REGION Network 96: "PALLET_PARA_ASCENSOR"
   RUNG wire#powerrail
      Contact( #Aux_1 )
      wire#w1
      Coil( "PALLET_PARA_ASCENSOR" )
   END_RUNG
   RUNG wire#powerrail
      Contact( "PALLET_PARA_ASCENSOR" )
      I_Contact( "Tonof_PALLET_EN_ASCENSOR" )
   END_RUNG wire#w1
   // the same network as SCL:
   "PALLET_PARA_ASCENSOR" := #Aux_1 OR ("PALLET_PARA_ASCENSOR" AND NOT "Tonof_PALLET_EN_ASCENSOR");
END_REGION

REGION Network 97: "PALLET_NO_FUERA_ASCENSOR" #Aux_1
   "IEC_Timer_0_DB_6".TOF(IN := NOT "iSnsPallEnAscen" AND NOT "iSnsSegAscenBajar", PT := T#500ms);
   #Aux_1 := "IEC_Timer_0_DB_6".Q;
END_REGION

REGION Network 98: "PALLET_NO_FUERA_ASCENSOR"
   RUNG wire#powerrail
      Contact( "iSnsPallEnAscen" )
      S_SR(operand := "PALLET_NO_FUERA_ASCENSOR", r1 := #Aux_1)
   END_RUNG
   // the same network as SCL:
   IF "iSnsPallEnAscen" THEN
       "PALLET_NO_FUERA_ASCENSOR" := TRUE;   // SR flip-flop
   END_IF;
   IF #Aux_1 THEN "PALLET_NO_FUERA_ASCENSOR" := FALSE; END_IF;
END_REGION

REGION Network 99: Aux PALLET_FUERA_TRANSP_2
   RUNG wire#powerrail
      Contact( "TRANSP_2_POR_ENVÍO" )
      Contact( "flanco".niSnsPallTrnsp_2 )
      S_SR(operand := #Aux_1, r1 := wire#w1)
   END_RUNG
   RUNG wire#powerrail
      Contact( "TRANSP_2_POR_RECAMBIO" )
      I_Contact( "TRANSP_2_POR_ENVÍO" )
   END_RUNG wire#w1
   // the same network as SCL:
   IF "TRANSP_2_POR_ENVÍO" AND "flanco".niSnsPallTrnsp_2 THEN
       #Aux_1 := TRUE;   // SR flip-flop
   END_IF;
   IF "TRANSP_2_POR_RECAMBIO" AND NOT "TRANSP_2_POR_ENVÍO" THEN #Aux_1 := FALSE; END_IF;
END_REGION

REGION Network 100: "PALLET_SALIO_TRANSP_2"
   "IEC_Timer_0_DB_9".TON(IN := #Aux_1, PT := T#1s);
   "PALLET_SALIO_TRANSP_2" := "IEC_Timer_0_DB_9".Q;
END_REGION

REGION Network 101: ZONA_ENVOLVEDORA_LIBRE
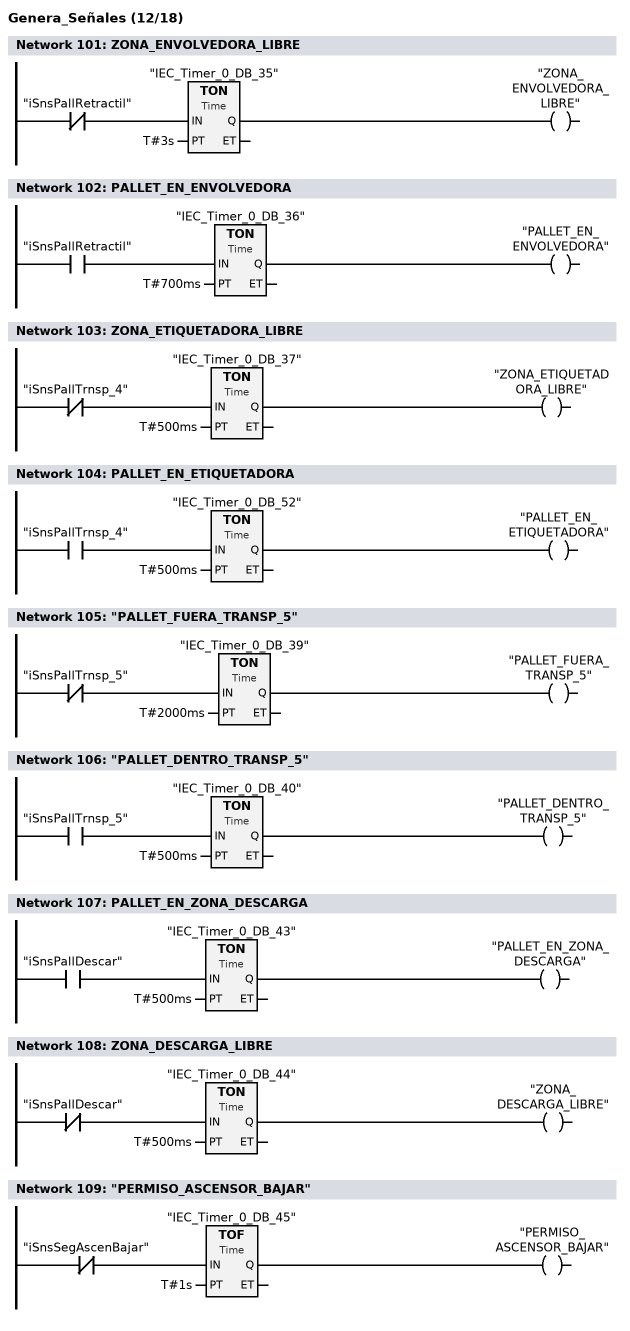
   "IEC_Timer_0_DB_35".TON(IN := NOT "iSnsPallRetractil", PT := T#3s);
   "ZONA_ENVOLVEDORA_LIBRE" := "IEC_Timer_0_DB_35".Q;
END_REGION

REGION Network 102: PALLET_EN_ENVOLVEDORA
   "IEC_Timer_0_DB_36".TON(IN := "iSnsPallRetractil", PT := T#700ms);
   "PALLET_EN_ENVOLVEDORA" := "IEC_Timer_0_DB_36".Q;
END_REGION

REGION Network 103: ZONA_ETIQUETADORA_LIBRE
   "IEC_Timer_0_DB_37".TON(IN := NOT "iSnsPallTrnsp_4", PT := T#500ms);
   "ZONA_ETIQUETADORA_LIBRE" := "IEC_Timer_0_DB_37".Q;
END_REGION

REGION Network 104: PALLET_EN_ETIQUETADORA
   "IEC_Timer_0_DB_52".TON(IN := "iSnsPallTrnsp_4", PT := T#500ms);
   "PALLET_EN_ETIQUETADORA" := "IEC_Timer_0_DB_52".Q;
END_REGION

REGION Network 105: "PALLET_FUERA_TRANSP_5"
   "IEC_Timer_0_DB_39".TON(IN := NOT "iSnsPallTrnsp_5", PT := T#2000ms);
   "PALLET_FUERA_TRANSP_5" := "IEC_Timer_0_DB_39".Q;
END_REGION

REGION Network 106: "PALLET_DENTRO_TRANSP_5"
   "IEC_Timer_0_DB_40".TON(IN := "iSnsPallTrnsp_5", PT := T#500ms);
   "PALLET_DENTRO_TRANSP_5" := "IEC_Timer_0_DB_40".Q;
END_REGION

REGION Network 107: PALLET_EN_ZONA_DESCARGA
   "IEC_Timer_0_DB_43".TON(IN := "iSnsPallDescar", PT := T#500ms);
   "PALLET_EN_ZONA_DESCARGA" := "IEC_Timer_0_DB_43".Q;
END_REGION

REGION Network 108: ZONA_DESCARGA_LIBRE
   "IEC_Timer_0_DB_44".TON(IN := NOT "iSnsPallDescar", PT := T#500ms);
   "ZONA_DESCARGA_LIBRE" := "IEC_Timer_0_DB_44".Q;
END_REGION

REGION Network 109: "PERMISO_ASCENSOR_BAJAR"
   "IEC_Timer_0_DB_45".TOF(IN := NOT "iSnsSegAscenBajar", PT := T#1s);
   "PERMISO_ASCENSOR_BAJAR" := "IEC_Timer_0_DB_45".Q;
END_REGION

REGION Network 110: "Pallet_Vacío_enPosición"
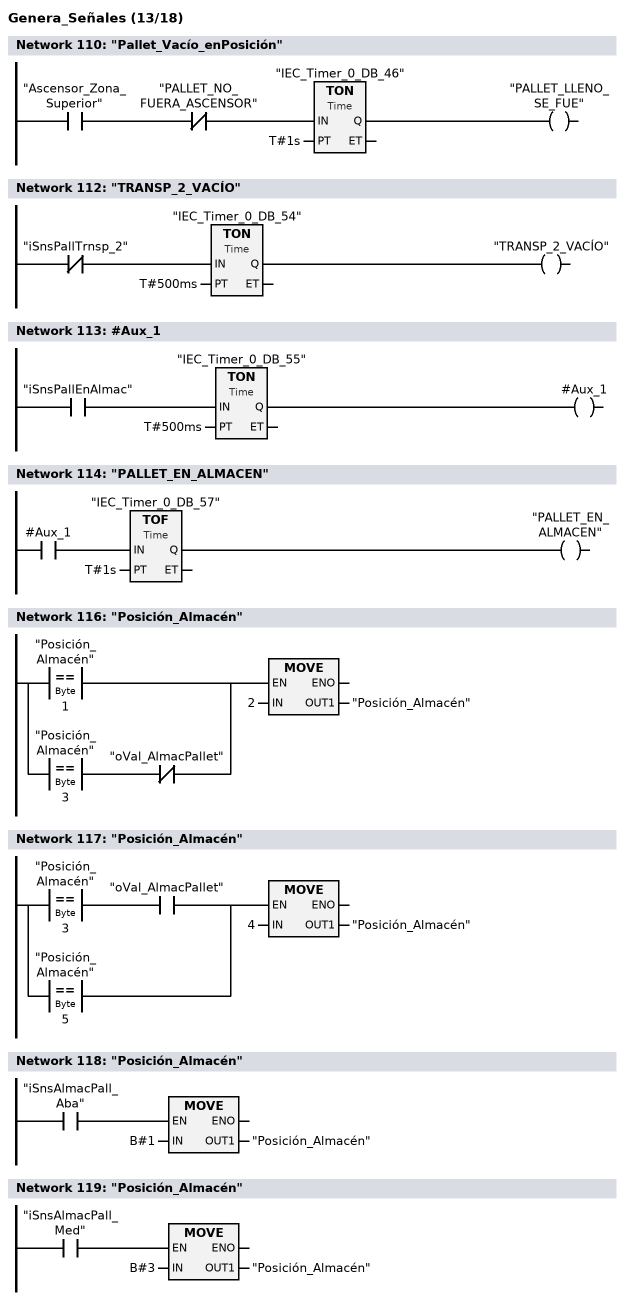
   "IEC_Timer_0_DB_46".TON(IN := "Ascensor_Zona_Superior" AND NOT "PALLET_NO_FUERA_ASCENSOR", PT := T#1s);
   "PALLET_LLENO_SE_FUE" := "IEC_Timer_0_DB_46".Q;
END_REGION

REGION Network 112: "TRANSP_2_VACÍO"
   "IEC_Timer_0_DB_54".TON(IN := NOT "iSnsPallTrnsp_2", PT := T#500ms);
   "TRANSP_2_VACÍO" := "IEC_Timer_0_DB_54".Q;
END_REGION

REGION Network 113: #Aux_1
   "IEC_Timer_0_DB_55".TON(IN := "iSnsPallEnAlmac", PT := T#500ms);
   #Aux_1 := "IEC_Timer_0_DB_55".Q;
END_REGION

REGION Network 114: "PALLET_EN_ALMACEN"
   "IEC_Timer_0_DB_57".TOF(IN := #Aux_1, PT := T#1s);
   "PALLET_EN_ALMACEN" := "IEC_Timer_0_DB_57".Q;
END_REGION

REGION Network 116: "Posición_Almacén"
   RUNG wire#powerrail
      { S7_Templates := "SrcType := Byte" } EQ_Contact(in1 := "Posición_Almacén", in2 := 1)
      wire#w1
      { S7_GenerateENO := "TRUE" } Move(in := 2, out1 => "Posición_Almacén")
   END_RUNG
   RUNG wire#powerrail
      { S7_Templates := "SrcType := Byte" } EQ_Contact(in1 := "Posición_Almacén", in2 := 3)
      I_Contact( "oVal_AlmacPallet" )
   END_RUNG wire#w1
   // the same network as SCL:
   IF ("Posición_Almacén" = 1) OR (("Posición_Almacén" = 3) AND NOT "oVal_AlmacPallet") THEN
       "Posición_Almacén" := 2;
   END_IF;
END_REGION

REGION Network 117: "Posición_Almacén"
   RUNG wire#powerrail
      { S7_Templates := "SrcType := Byte" } EQ_Contact(in1 := "Posición_Almacén", in2 := 3)
      Contact( "oVal_AlmacPallet" )
      wire#w1
      { S7_GenerateENO := "TRUE" } Move(in := 4, out1 => "Posición_Almacén")
   END_RUNG
   RUNG wire#powerrail
      { S7_Templates := "SrcType := Byte" } EQ_Contact(in1 := "Posición_Almacén", in2 := 5)
   END_RUNG wire#w1
   // the same network as SCL:
   IF (("Posición_Almacén" = 3) AND "oVal_AlmacPallet") OR ("Posición_Almacén" = 5) THEN
       "Posición_Almacén" := 4;
   END_IF;
END_REGION

REGION Network 118: "Posición_Almacén"
   RUNG wire#powerrail
      Contact( "iSnsAlmacPall_Aba" )
      { S7_GenerateENO := "TRUE" } Move(in := B#1, out1 => "Posición_Almacén")
   END_RUNG
   // the same network as SCL:
   IF "iSnsAlmacPall_Aba" THEN "Posición_Almacén" := B#1; END_IF;
END_REGION

REGION Network 119: "Posición_Almacén"
   RUNG wire#powerrail
      Contact( "iSnsAlmacPall_Med" )
      { S7_GenerateENO := "TRUE" } Move(in := B#3, out1 => "Posición_Almacén")
   END_RUNG
   // the same network as SCL:
   IF "iSnsAlmacPall_Med" THEN "Posición_Almacén" := B#3; END_IF;
END_REGION

REGION Network 120: "Posición_Almacén"
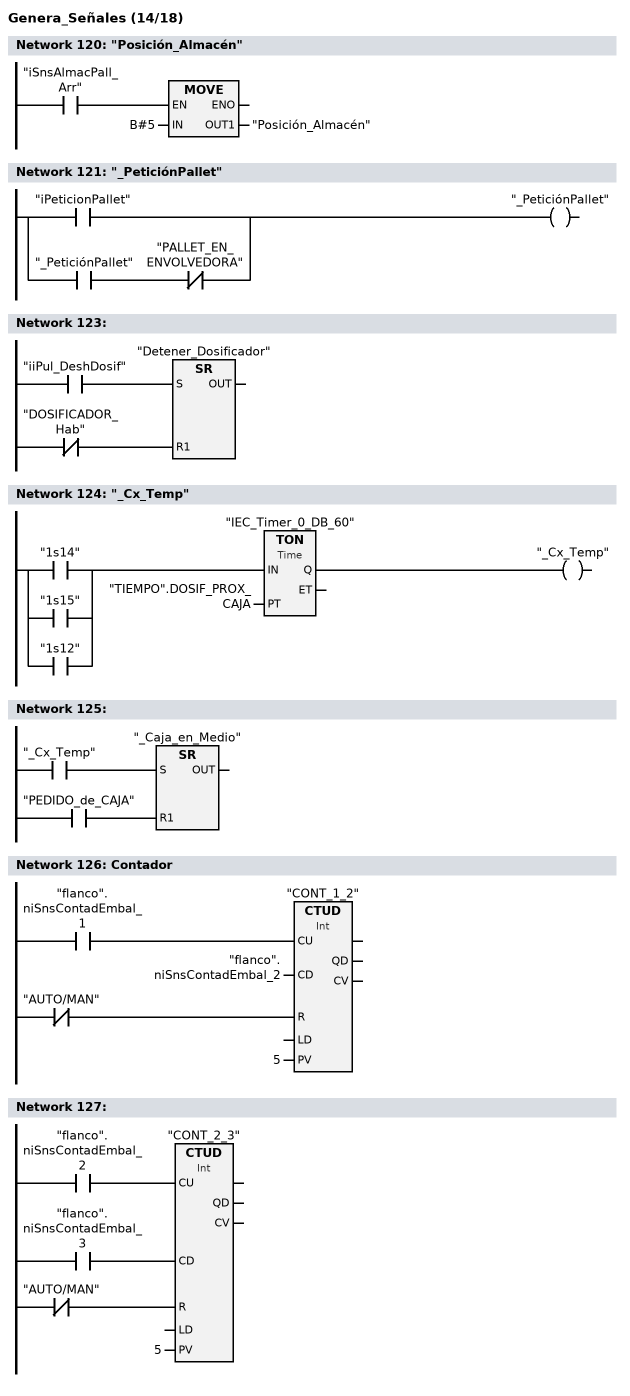
   RUNG wire#powerrail
      Contact( "iSnsAlmacPall_Arr" )
      { S7_GenerateENO := "TRUE" } Move(in := B#5, out1 => "Posición_Almacén")
   END_RUNG
   // the same network as SCL:
   IF "iSnsAlmacPall_Arr" THEN "Posición_Almacén" := B#5; END_IF;
END_REGION

REGION Network 121: "_PeticiónPallet"
   RUNG wire#powerrail
      Contact( "iPeticionPallet" )
      wire#w1
      Coil( "_PeticiónPallet" )
   END_RUNG
   RUNG wire#powerrail
      Contact( "_PeticiónPallet" )
      I_Contact( "PALLET_EN_ENVOLVEDORA" )
   END_RUNG wire#w1
   // the same network as SCL:
   "_PeticiónPallet" := "iPeticionPallet" OR ("_PeticiónPallet" AND NOT "PALLET_EN_ENVOLVEDORA");
END_REGION

REGION Network 122: ----------------------------------------------------------------------- DOSIFICADOR ---------------------------------------------------------------------------
END_REGION

REGION Network 123
   RUNG wire#powerrail
      Contact( "iiPul_DeshDosif" )
      S_SR(operand := "Detener_Dosificador", r1 := wire#w1)
   END_RUNG
   RUNG wire#powerrail
      I_Contact( "DOSIFICADOR_Hab" )
   END_RUNG wire#w1
   // the same network as SCL:
   IF "iiPul_DeshDosif" THEN
       "Detener_Dosificador" := TRUE;   // SR flip-flop
   END_IF;
   IF NOT "DOSIFICADOR_Hab" THEN "Detener_Dosificador" := FALSE; END_IF;
END_REGION

REGION Network 124: "_Cx_Temp"
   "IEC_Timer_0_DB_60".TON(IN := "1s14" OR "1s15" OR "1s12", PT := "TIEMPO".DOSIF_PROX_CAJA);
   "_Cx_Temp" := "IEC_Timer_0_DB_60".Q;
END_REGION

REGION Network 125
   RUNG wire#powerrail
      Contact( "_Cx_Temp" )
      S_SR(operand := "_Caja_en_Medio", r1 := wire#w1)
   END_RUNG
   RUNG wire#powerrail
      Contact( "PEDIDO_de_CAJA" )
   END_RUNG wire#w1
   // the same network as SCL:
   IF "_Cx_Temp" THEN
       "_Caja_en_Medio" := TRUE;   // SR flip-flop
   END_IF;
   IF "PEDIDO_de_CAJA" THEN "_Caja_en_Medio" := FALSE; END_IF;
END_REGION

REGION Network 126: Contador
   "CONT_1_2".CTUD(CU := "flanco".niSnsContadEmbal_1,
                   CD := "flanco".niSnsContadEmbal_2,
                   R := NOT "AUTO/MAN",
                   PV := 5);
END_REGION

REGION Network 127
   "CONT_2_3".CTUD(CU := "flanco".niSnsContadEmbal_2,
                   CD := "flanco".niSnsContadEmbal_3,
                   R := NOT "AUTO/MAN",
                   PV := 5);
END_REGION

REGION Network 129: SET "Anterior_Vertical"
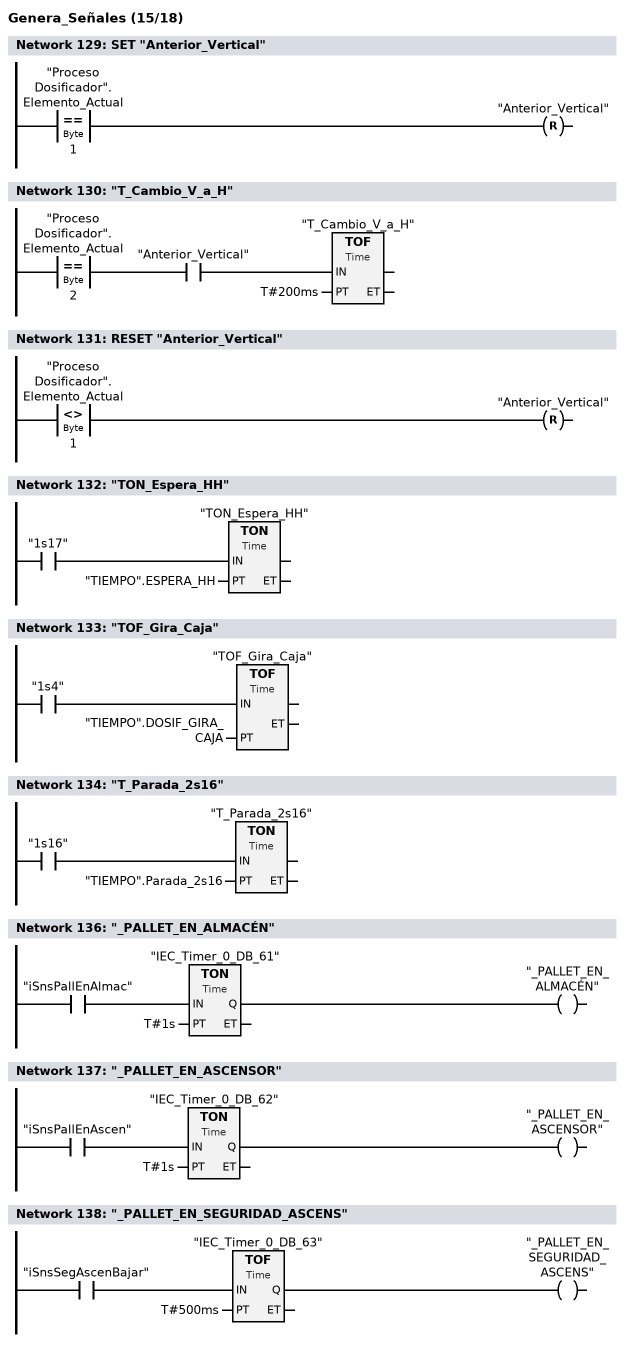
   RUNG wire#powerrail
      { S7_Templates := "SrcType := Byte" } EQ_Contact(in1 := "Proceso Dosificador".Elemento_Actual, in2 := 1)
      R_Coil( "Anterior_Vertical" )
   END_RUNG
   // the same network as SCL:
   IF "Proceso Dosificador".Elemento_Actual = 1 THEN "Anterior_Vertical" := FALSE; END_IF;
END_REGION

REGION Network 130: "T_Cambio_V_a_H"
   "T_Cambio_V_a_H".TOF(IN := ("Proceso Dosificador".Elemento_Actual = 2) AND "Anterior_Vertical",
                        PT := T#200ms);
END_REGION

REGION Network 131: RESET "Anterior_Vertical"
   RUNG wire#powerrail
      { S7_Templates := "SrcType := Byte" } NE_Contact(in1 := "Proceso Dosificador".Elemento_Actual, in2 := 1)
      R_Coil( "Anterior_Vertical" )
   END_RUNG
   // the same network as SCL:
   IF "Proceso Dosificador".Elemento_Actual <> 1 THEN "Anterior_Vertical" := FALSE; END_IF;
END_REGION

REGION Network 132: "TON_Espera_HH"
   "TON_Espera_HH".TON(IN := "1s17", PT := "TIEMPO".ESPERA_HH);
END_REGION

REGION Network 133: "TOF_Gira_Caja"
   "TOF_Gira_Caja".TOF(IN := "1s4", PT := "TIEMPO".DOSIF_GIRA_CAJA);
END_REGION

REGION Network 134: "T_Parada_2s16"
   "T_Parada_2s16".TON(IN := "1s16", PT := "TIEMPO".Parada_2s16);
END_REGION

REGION Network 135: ----------------------------------------------------------------------- TRANSPORTE PALLETS 2 ---------------------------------------------------------------------------
END_REGION

REGION Network 136: "_PALLET_EN_ALMACÉN"
   "IEC_Timer_0_DB_61".TON(IN := "iSnsPallEnAlmac", PT := T#1s);
   "_PALLET_EN_ALMACÉN" := "IEC_Timer_0_DB_61".Q;
END_REGION

REGION Network 137: "_PALLET_EN_ASCENSOR"
   "IEC_Timer_0_DB_62".TON(IN := "iSnsPallEnAscen", PT := T#1s);
   "_PALLET_EN_ASCENSOR" := "IEC_Timer_0_DB_62".Q;
END_REGION

REGION Network 138: "_PALLET_EN_SEGURIDAD_ASCENS"
   "IEC_Timer_0_DB_63".TOF(IN := "iSnsSegAscenBajar", PT := T#500ms);
   "_PALLET_EN_SEGURIDAD_ASCENS" := "IEC_Timer_0_DB_63".Q;
END_REGION

REGION Network 139: "_PALLET_EN_TRANSP_2"
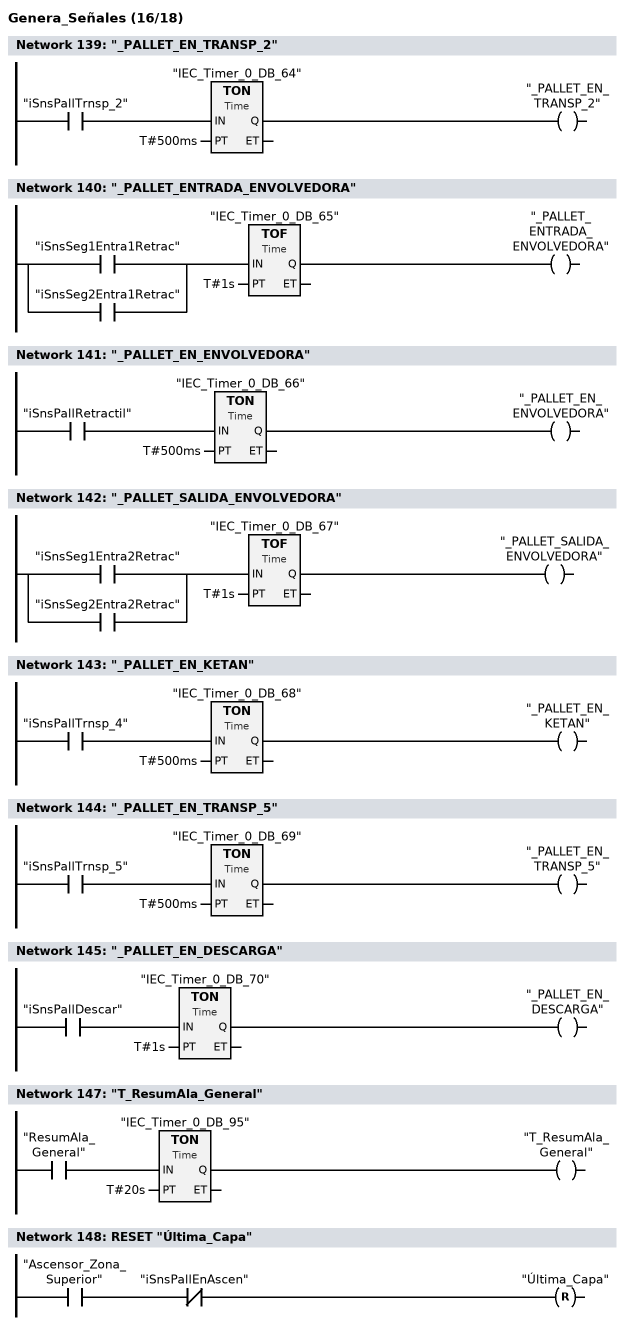
   "IEC_Timer_0_DB_64".TON(IN := "iSnsPallTrnsp_2", PT := T#500ms);
   "_PALLET_EN_TRANSP_2" := "IEC_Timer_0_DB_64".Q;
END_REGION

REGION Network 140: "_PALLET_ENTRADA_ENVOLVEDORA"
   "IEC_Timer_0_DB_65".TOF(IN := "iSnsSeg1Entra1Retrac" OR "iSnsSeg2Entra1Retrac", PT := T#1s);
   "_PALLET_ENTRADA_ENVOLVEDORA" := "IEC_Timer_0_DB_65".Q;
END_REGION

REGION Network 141: "_PALLET_EN_ENVOLVEDORA"
   "IEC_Timer_0_DB_66".TON(IN := "iSnsPallRetractil", PT := T#500ms);
   "_PALLET_EN_ENVOLVEDORA" := "IEC_Timer_0_DB_66".Q;
END_REGION

REGION Network 142: "_PALLET_SALIDA_ENVOLVEDORA"
   "IEC_Timer_0_DB_67".TOF(IN := "iSnsSeg1Entra2Retrac" OR "iSnsSeg2Entra2Retrac", PT := T#1s);
   "_PALLET_SALIDA_ENVOLVEDORA" := "IEC_Timer_0_DB_67".Q;
END_REGION

REGION Network 143: "_PALLET_EN_KETAN"
   "IEC_Timer_0_DB_68".TON(IN := "iSnsPallTrnsp_4", PT := T#500ms);
   "_PALLET_EN_KETAN" := "IEC_Timer_0_DB_68".Q;
END_REGION

REGION Network 144: "_PALLET_EN_TRANSP_5"
   "IEC_Timer_0_DB_69".TON(IN := "iSnsPallTrnsp_5", PT := T#500ms);
   "_PALLET_EN_TRANSP_5" := "IEC_Timer_0_DB_69".Q;
END_REGION

REGION Network 145: "_PALLET_EN_DESCARGA"
   "IEC_Timer_0_DB_70".TON(IN := "iSnsPallDescar", PT := T#1s);
   "_PALLET_EN_DESCARGA" := "IEC_Timer_0_DB_70".Q;
END_REGION

REGION Network 146: ----------------------------------------------------------------------- GENERAL ---------------------------------------------------------------------------
END_REGION

REGION Network 147: "T_ResumAla_General"
   "IEC_Timer_0_DB_95".TON(IN := "ResumAla_General", PT := T#20s);
   "T_ResumAla_General" := "IEC_Timer_0_DB_95".Q;
END_REGION

REGION Network 148: RESET "Última_Capa"
   RUNG wire#powerrail
      Contact( "Ascensor_Zona_Superior" )
      I_Contact( "iSnsPallEnAscen" )
      R_Coil( "Última_Capa" )
   END_RUNG
   // the same network as SCL:
   IF "Ascensor_Zona_Superior" AND NOT "iSnsPallEnAscen" THEN "Última_Capa" := FALSE; END_IF;
END_REGION

REGION Network 149: "Tag_2" se activa si el ascensor baja con la señal "Última_Capa" activada
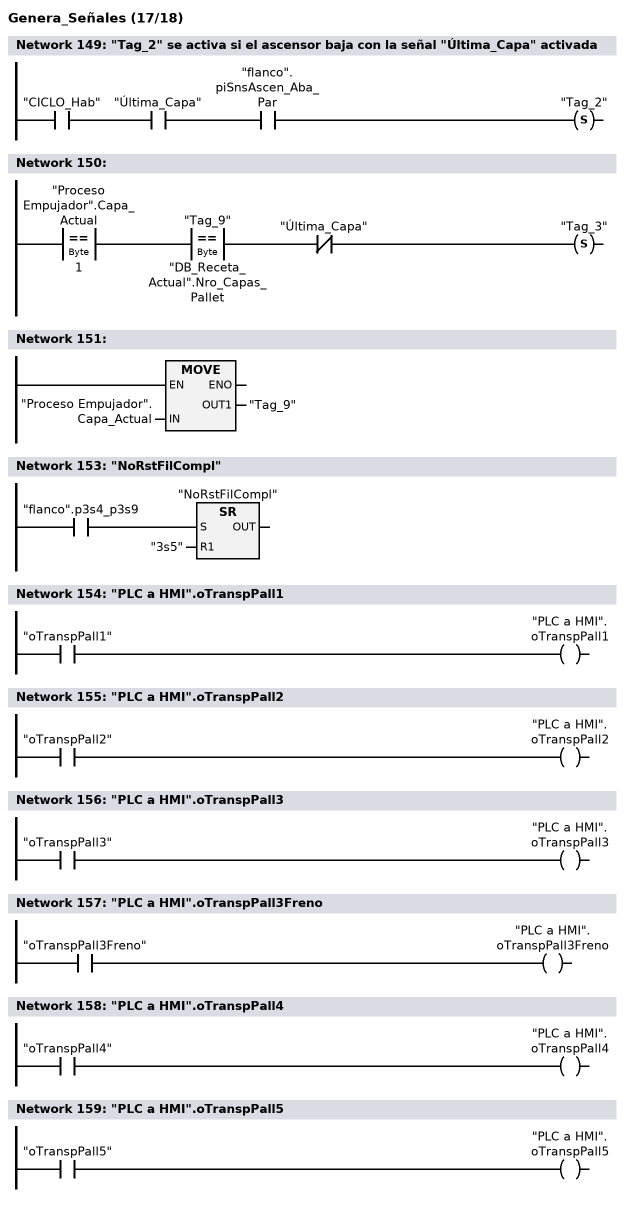
   RUNG wire#powerrail
      Contact( "CICLO_Hab" )
      Contact( "Última_Capa" )
      Contact( "flanco".piSnsAscen_Aba_Par )
      S_Coil( "Tag_2" )
   END_RUNG
   // the same network as SCL:
   IF "CICLO_Hab" AND "Última_Capa" AND "flanco".piSnsAscen_Aba_Par THEN "Tag_2" := TRUE; END_IF;
END_REGION

REGION Network 150
   RUNG wire#powerrail
      { S7_Templates := "SrcType := Byte" } EQ_Contact(in1 := "Proceso Empujador".Capa_Actual, in2 := 1)
      { S7_Templates := "SrcType := Byte" } EQ_Contact(in1 := "Tag_9", in2 := "DB_Receta_Actual".Nro_Capas_Pallet)
      I_Contact( "Última_Capa" )
      S_Coil( "Tag_3" )
   END_RUNG
   // the same network as SCL:
   IF ("Proceso Empujador".Capa_Actual = 1) AND ("Tag_9" = "DB_Receta_Actual".Nro_Capas_Pallet) AND NOT "Última_Capa" THEN
       "Tag_3" := TRUE;
   END_IF;
END_REGION

REGION Network 151
   RUNG wire#powerrail
      { S7_GenerateENO := "TRUE" } Move(in := "Proceso Empujador".Capa_Actual, out1 => "Tag_9")
   END_RUNG
   // the same network as SCL:
   "Tag_9" := "Proceso Empujador".Capa_Actual;
END_REGION

REGION Network 152 (STL): en AWL se inrementa un Byte
         A     "flanco"."pHMI.Pls_Inc_Figura_Sel";
         JCN   fin;
         L     "DB_Animación".Figura_SEL;
         INC   1;
         T     "DB_Animación".Figura_SEL;
   fin:  NOP   0;
END_REGION

REGION Network 153: "NoRstFilCompl"
   RUNG wire#powerrail
      Contact( "flanco".p3s4_p3s9 )
      S_SR(operand := "NoRstFilCompl", r1 := "3s5")
   END_RUNG
   // the same network as SCL:
   IF "flanco".p3s4_p3s9 THEN
       "NoRstFilCompl" := TRUE;   // SR flip-flop
   END_IF;
   IF "3s5" THEN "NoRstFilCompl" := FALSE; END_IF;
END_REGION

REGION Network 154: "PLC a HMI".oTranspPall1
   RUNG wire#powerrail
      Contact( "oTranspPall1" )
      Coil( "PLC a HMI".oTranspPall1 )
   END_RUNG
   // the same network as SCL:
   "PLC a HMI".oTranspPall1 := "oTranspPall1";
END_REGION

REGION Network 155: "PLC a HMI".oTranspPall2
   RUNG wire#powerrail
      Contact( "oTranspPall2" )
      Coil( "PLC a HMI".oTranspPall2 )
   END_RUNG
   // the same network as SCL:
   "PLC a HMI".oTranspPall2 := "oTranspPall2";
END_REGION

REGION Network 156: "PLC a HMI".oTranspPall3
   RUNG wire#powerrail
      Contact( "oTranspPall3" )
      Coil( "PLC a HMI".oTranspPall3 )
   END_RUNG
   // the same network as SCL:
   "PLC a HMI".oTranspPall3 := "oTranspPall3";
END_REGION

REGION Network 157: "PLC a HMI".oTranspPall3Freno
   RUNG wire#powerrail
      Contact( "oTranspPall3Freno" )
      Coil( "PLC a HMI".oTranspPall3Freno )
   END_RUNG
   // the same network as SCL:
   "PLC a HMI".oTranspPall3Freno := "oTranspPall3Freno";
END_REGION

REGION Network 158: "PLC a HMI".oTranspPall4
   RUNG wire#powerrail
      Contact( "oTranspPall4" )
      Coil( "PLC a HMI".oTranspPall4 )
   END_RUNG
   // the same network as SCL:
   "PLC a HMI".oTranspPall4 := "oTranspPall4";
END_REGION

REGION Network 159: "PLC a HMI".oTranspPall5
   RUNG wire#powerrail
      Contact( "oTranspPall5" )
      Coil( "PLC a HMI".oTranspPall5 )
   END_RUNG
   // the same network as SCL:
   "PLC a HMI".oTranspPall5 := "oTranspPall5";
END_REGION

REGION Network 160: "Remanente".Set_para_2c13
   // En el estado 2s12 se espera a que se vaya el pallet lleno, una vez  llegado al estado 2s13 la señal pierde validez.
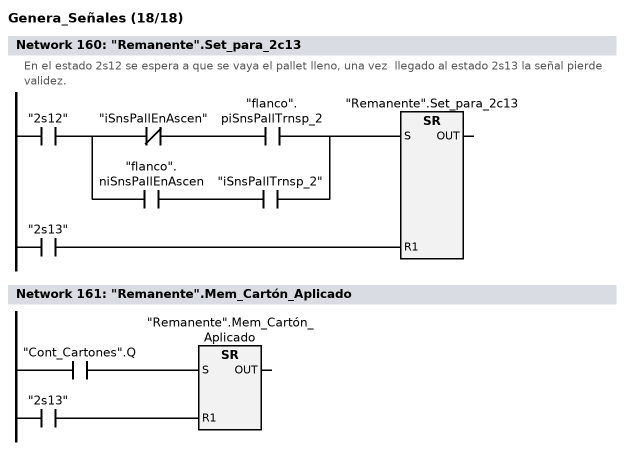
   RUNG wire#powerrail
      Contact( "2s12" )
      wire#w1
      I_Contact( "iSnsPallEnAscen" )
      Contact( "flanco".piSnsPallTrnsp_2 )
      wire#w2
      S_SR(operand := "Remanente".Set_para_2c13, r1 := wire#w3)
   END_RUNG
   RUNG wire#w1
      Contact( "flanco".niSnsPallEnAscen )
      Contact( "iSnsPallTrnsp_2" )
   END_RUNG wire#w2
   RUNG wire#powerrail
      Contact( "2s13" )
   END_RUNG wire#w3
   // the same network as SCL:
   IF "2s12" AND ((NOT "iSnsPallEnAscen" AND "flanco".piSnsPallTrnsp_2) OR ("flanco".niSnsPallEnAscen AND "iSnsPallTrnsp_2")) THEN
       "Remanente".Set_para_2c13 := TRUE;   // SR flip-flop
   END_IF;
   IF "2s13" THEN "Remanente".Set_para_2c13 := FALSE; END_IF;
END_REGION

REGION Network 161: "Remanente".Mem_Cartón_Aplicado
   RUNG wire#powerrail
      Contact( "Cont_Cartones".Q )
      S_SR(operand := "Remanente".Mem_Cartón_Aplicado, r1 := wire#w1)
   END_RUNG
   RUNG wire#powerrail
      Contact( "2s13" )
   END_RUNG wire#w1
   // the same network as SCL:
   IF "Cont_Cartones".Q THEN
       "Remanente".Mem_Cartón_Aplicado := TRUE;   // SR flip-flop
   END_IF;
   IF "2s13" THEN "Remanente".Mem_Cartón_Aplicado := FALSE; END_IF;
END_REGION
END_FUNCTION

FUNCTION "Activa_Pistón" : Void   // FC20, STL
{ S7_Optimized_Access := 'FALSE' }
VERSION : 0.1
BEGIN

REGION Network 1: Constantes
         L     38;
         T     #Length_Capas;
         L     54;
         T     #Offset_Capas;
END_REGION

REGION Network 2
         CLR;
         =     "Poner_Pistón";
END_REGION

REGION Network 3: #Adress_Capa
         L     1;
         L     "Proceso CargaPallet".Capa_Actual;
         <=I;
         JCN   Fin;
         DEC   1;
         L     #Length_Capas;
         *I;
         L     #Offset_Capas;
         +I;
         T     #Adress_Capa;
END_REGION

REGION Network 4: LAR1
         L     #Adress_Capa;
         L     36;  // Offset Usar Pistón
         +I;
         SLD   3;
         LAR1;
END_REGION

REGION Network 5: "Poner_Pistón"
         OPN   "DB_Receta_Actual";
         A     DBX [ AR1 , P#0.0 ];
         =     "Poner_Pistón";
   Fin:  NOP   0;
END_REGION
END_FUNCTION

FUNCTION "Conteo_MAN" : Void   // FC24, STL
{ S7_Optimized_Access := 'FALSE' }
VERSION : 0.1
BEGIN

REGION Network 1: Inc/Dec Capa
         L     "DB_Receta_Actual".Nro_Capas_Pallet;
         L     "Proceso Empujador".Capa_Actual;
         >I;
         =     #Habil_Inc;
         L     1;
         >I;
         =     #Habil_Dec;
         A     #Habil_Inc;
         A     "flanco"."nHMI.Pls_Inc_Capa";
         JCN   noInc;
         L     "Proceso Empujador".Capa_Actual;
         INC   1;
         T     "Proceso Empujador".Capa_Actual;
   noInc:A     #Habil_Dec;
         A     "flanco"."nHMI.Pls_Dec_Capa";
         JCN   noDec;
         L     "Proceso Empujador".Capa_Actual;
         DEC   1;
         T     "Proceso Empujador".Capa_Actual;
   noDec:NOP   0;

         A     "HMI".Pls_ResetPallets;
         JCN   noRePall;
         L     0;
         T     "Proceso Empujador".Cant_Pallets;
         T     "Proceso CargaPallet".Cant_Pallets;
   noRePall:NOP   0;
END_REGION

REGION Network 2
         L     "Proceso Empujador".Capa_Actual;
         DEC   1;
         T     "Proceso CargaPallet".Capa_Actual;
END_REGION
END_FUNCTION

FUNCTION "Interfase" : Void   // FC25, LAD
{ S7_Optimized_Access := 'FALSE' }
VERSION : 0.1
BEGIN

REGION Network 1: ------------------------------------------------------ ENVOLVEDORA STORK --------------------------------------------------------------
END_REGION

REGION Network 2: "oRetractiSeg"
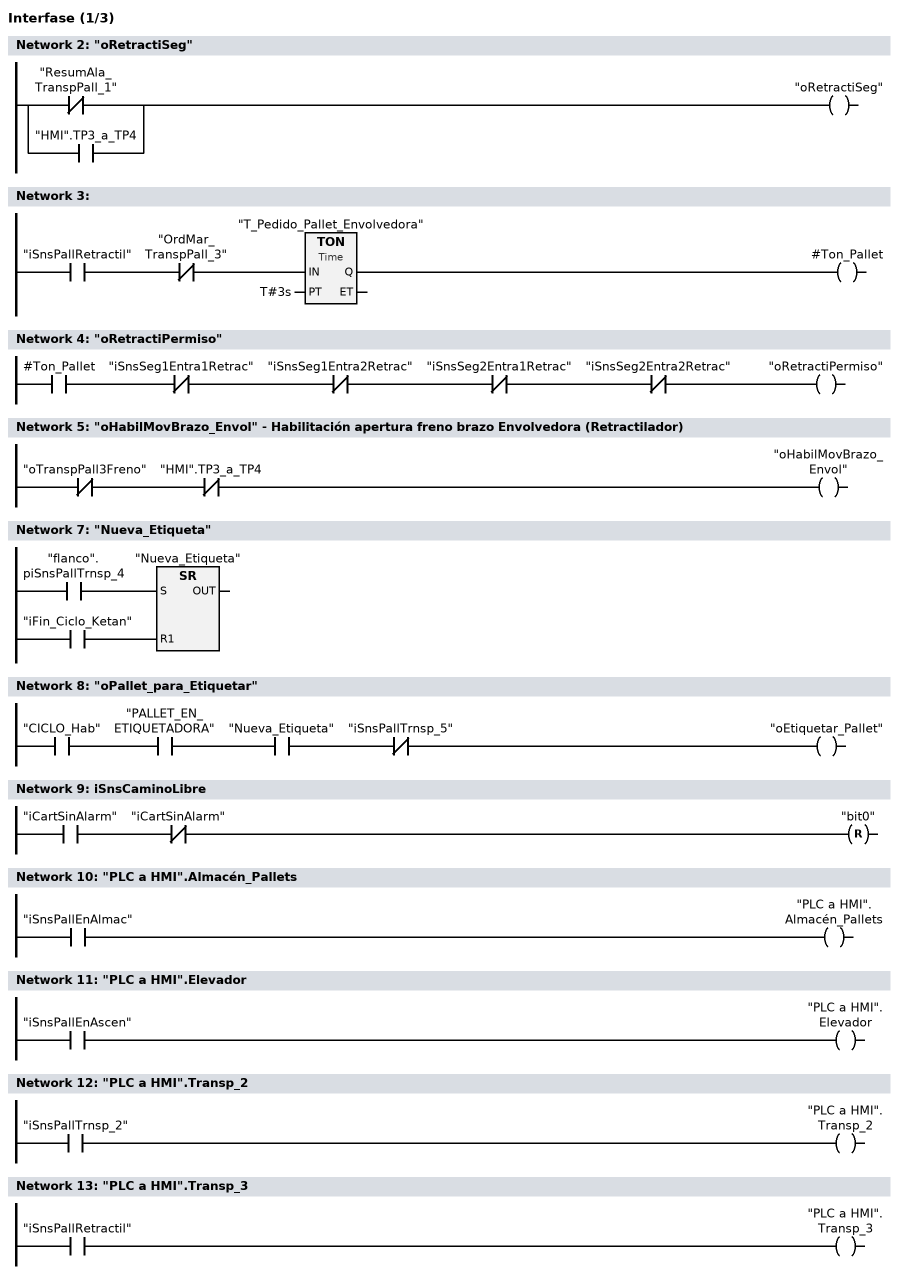
   RUNG wire#powerrail
      I_Contact( "ResumAla_TranspPall_1" )
      wire#w1
      Coil( "oRetractiSeg" )
   END_RUNG
   RUNG wire#powerrail
      Contact( "HMI".TP3_a_TP4 )
   END_RUNG wire#w1
   // the same network as SCL:
   "oRetractiSeg" := NOT "ResumAla_TranspPall_1" OR "HMI".TP3_a_TP4;
END_REGION

REGION Network 3
   "T_Pedido_Pallet_Envolvedora".TON(in := "iSnsPallRetractil" AND NOT "OrdMar_TranspPall_3", pt := T#3s);
   #Ton_Pallet := "T_Pedido_Pallet_Envolvedora".q;
END_REGION

REGION Network 4: "oRetractiPermiso"
   RUNG wire#powerrail
      Contact( #Ton_Pallet )
      I_Contact( "iSnsSeg1Entra1Retrac" )
      I_Contact( "iSnsSeg1Entra2Retrac" )
      I_Contact( "iSnsSeg2Entra1Retrac" )
      I_Contact( "iSnsSeg2Entra2Retrac" )
      Coil( "oRetractiPermiso" )
   END_RUNG
   // the same network as SCL:
   "oRetractiPermiso" := #Ton_Pallet AND NOT "iSnsSeg1Entra1Retrac" AND NOT "iSnsSeg1Entra2Retrac" AND NOT "iSnsSeg2Entra1Retrac" AND NOT "iSnsSeg2Entra2Retrac";
END_REGION

REGION Network 5: "oHabilMovBrazo_Envol" - Habilitación apertura freno brazo Envolvedora (Retractilador)
   RUNG wire#powerrail
      I_Contact( "oTranspPall3Freno" )
      I_Contact( "HMI".TP3_a_TP4 )
      Coil( "oHabilMovBrazo_Envol" )
   END_RUNG
   // the same network as SCL:
   "oHabilMovBrazo_Envol" := NOT "oTranspPall3Freno" AND NOT "HMI".TP3_a_TP4;
END_REGION

REGION Network 6: ------------------------------------------------------ ETIQUETADORA KETAN --------------------------------------------------------------
END_REGION

REGION Network 7: "Nueva_Etiqueta"
   RUNG wire#powerrail
      Contact( "flanco".piSnsPallTrnsp_4 )
      S_SR(operand := "Nueva_Etiqueta", r1 := wire#w1)
   END_RUNG
   RUNG wire#powerrail
      Contact( "iFin_Ciclo_Ketan" )
   END_RUNG wire#w1
   // the same network as SCL:
   IF "flanco".piSnsPallTrnsp_4 THEN
       "Nueva_Etiqueta" := TRUE;   // SR flip-flop
   END_IF;
   IF "iFin_Ciclo_Ketan" THEN "Nueva_Etiqueta" := FALSE; END_IF;
END_REGION

REGION Network 8: "oPallet_para_Etiquetar"
   RUNG wire#powerrail
      Contact( "CICLO_Hab" )
      Contact( "PALLET_EN_ETIQUETADORA" )
      Contact( "Nueva_Etiqueta" )
      I_Contact( "iSnsPallTrnsp_5" )
      Coil( "oEtiquetar_Pallet" )
   END_RUNG
   // the same network as SCL:
   "oEtiquetar_Pallet" := "CICLO_Hab" AND "PALLET_EN_ETIQUETADORA" AND "Nueva_Etiqueta" AND NOT "iSnsPallTrnsp_5";
END_REGION

REGION Network 9: iSnsCaminoLibre
   RUNG wire#powerrail
      Contact( "iCartSinAlarm" )
      I_Contact( "iCartSinAlarm" )
      R_Coil( "bit0" )
   END_RUNG
   // the same network as SCL:
   IF "iCartSinAlarm" AND NOT "iCartSinAlarm" THEN "bit0" := FALSE; END_IF;
END_REGION

REGION Network 10: "PLC a HMI".Almacén_Pallets
   RUNG wire#powerrail
      Contact( "iSnsPallEnAlmac" )
      Coil( "PLC a HMI".Almacén_Pallets )
   END_RUNG
   // the same network as SCL:
   "PLC a HMI".Almacén_Pallets := "iSnsPallEnAlmac";
END_REGION

REGION Network 11: "PLC a HMI".Elevador
   RUNG wire#powerrail
      Contact( "iSnsPallEnAscen" )
      Coil( "PLC a HMI".Elevador )
   END_RUNG
   // the same network as SCL:
   "PLC a HMI".Elevador := "iSnsPallEnAscen";
END_REGION

REGION Network 12: "PLC a HMI".Transp_2
   RUNG wire#powerrail
      Contact( "iSnsPallTrnsp_2" )
      Coil( "PLC a HMI".Transp_2 )
   END_RUNG
   // the same network as SCL:
   "PLC a HMI".Transp_2 := "iSnsPallTrnsp_2";
END_REGION

REGION Network 13: "PLC a HMI".Transp_3
   RUNG wire#powerrail
      Contact( "iSnsPallRetractil" )
      Coil( "PLC a HMI".Transp_3 )
   END_RUNG
   // the same network as SCL:
   "PLC a HMI".Transp_3 := "iSnsPallRetractil";
END_REGION

REGION Network 14: "PLC a HMI".Transp_4
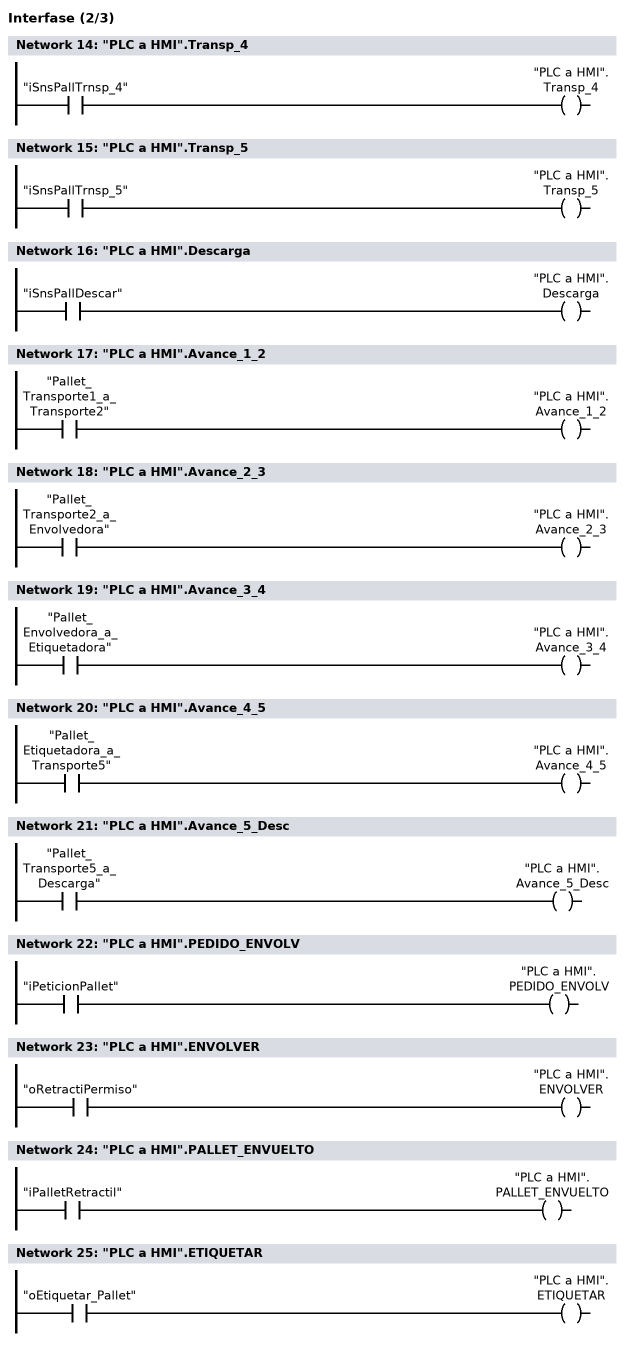
   RUNG wire#powerrail
      Contact( "iSnsPallTrnsp_4" )
      Coil( "PLC a HMI".Transp_4 )
   END_RUNG
   // the same network as SCL:
   "PLC a HMI".Transp_4 := "iSnsPallTrnsp_4";
END_REGION

REGION Network 15: "PLC a HMI".Transp_5
   RUNG wire#powerrail
      Contact( "iSnsPallTrnsp_5" )
      Coil( "PLC a HMI".Transp_5 )
   END_RUNG
   // the same network as SCL:
   "PLC a HMI".Transp_5 := "iSnsPallTrnsp_5";
END_REGION

REGION Network 16: "PLC a HMI".Descarga
   RUNG wire#powerrail
      Contact( "iSnsPallDescar" )
      Coil( "PLC a HMI".Descarga )
   END_RUNG
   // the same network as SCL:
   "PLC a HMI".Descarga := "iSnsPallDescar";
END_REGION

REGION Network 17: "PLC a HMI".Avance_1_2
   RUNG wire#powerrail
      Contact( "Pallet_Transporte1_a_Transporte2" )
      Coil( "PLC a HMI".Avance_1_2 )
   END_RUNG
   // the same network as SCL:
   "PLC a HMI".Avance_1_2 := "Pallet_Transporte1_a_Transporte2";
END_REGION

REGION Network 18: "PLC a HMI".Avance_2_3
   RUNG wire#powerrail
      Contact( "Pallet_Transporte2_a_Envolvedora" )
      Coil( "PLC a HMI".Avance_2_3 )
   END_RUNG
   // the same network as SCL:
   "PLC a HMI".Avance_2_3 := "Pallet_Transporte2_a_Envolvedora";
END_REGION

REGION Network 19: "PLC a HMI".Avance_3_4
   RUNG wire#powerrail
      Contact( "Pallet_Envolvedora_a_Etiquetadora" )
      Coil( "PLC a HMI".Avance_3_4 )
   END_RUNG
   // the same network as SCL:
   "PLC a HMI".Avance_3_4 := "Pallet_Envolvedora_a_Etiquetadora";
END_REGION

REGION Network 20: "PLC a HMI".Avance_4_5
   RUNG wire#powerrail
      Contact( "Pallet_Etiquetadora_a_Transporte5" )
      Coil( "PLC a HMI".Avance_4_5 )
   END_RUNG
   // the same network as SCL:
   "PLC a HMI".Avance_4_5 := "Pallet_Etiquetadora_a_Transporte5";
END_REGION

REGION Network 21: "PLC a HMI".Avance_5_Desc
   RUNG wire#powerrail
      Contact( "Pallet_Transporte5_a_Descarga" )
      Coil( "PLC a HMI".Avance_5_Desc )
   END_RUNG
   // the same network as SCL:
   "PLC a HMI".Avance_5_Desc := "Pallet_Transporte5_a_Descarga";
END_REGION

REGION Network 22: "PLC a HMI".PEDIDO_ENVOLV
   RUNG wire#powerrail
      Contact( "iPeticionPallet" )
      Coil( "PLC a HMI".PEDIDO_ENVOLV )
   END_RUNG
   // the same network as SCL:
   "PLC a HMI".PEDIDO_ENVOLV := "iPeticionPallet";
END_REGION

REGION Network 23: "PLC a HMI".ENVOLVER
   RUNG wire#powerrail
      Contact( "oRetractiPermiso" )
      Coil( "PLC a HMI".ENVOLVER )
   END_RUNG
   // the same network as SCL:
   "PLC a HMI".ENVOLVER := "oRetractiPermiso";
END_REGION

REGION Network 24: "PLC a HMI".PALLET_ENVUELTO
   RUNG wire#powerrail
      Contact( "iPalletRetractil" )
      Coil( "PLC a HMI".PALLET_ENVUELTO )
   END_RUNG
   // the same network as SCL:
   "PLC a HMI".PALLET_ENVUELTO := "iPalletRetractil";
END_REGION

REGION Network 25: "PLC a HMI".ETIQUETAR
   RUNG wire#powerrail
      Contact( "oEtiquetar_Pallet" )
      Coil( "PLC a HMI".ETIQUETAR )
   END_RUNG
   // the same network as SCL:
   "PLC a HMI".ETIQUETAR := "oEtiquetar_Pallet";
END_REGION

REGION Network 26: "PLC a HMI".CICLO_OK
